(* Logix 5000 project; controller PLC_MCC1300_75F1 vendor 1 type 14 code 166 rev 32.11; software revision 32.04; part 2 of 83 *)

TYPE MAC_Popup_ZC_ALM :
STRUCT
   rgxStoppingFault : DINT[1];   // Generic stopping faults
   rgxFault : DINT[1];   // Generic faults
   rgxWarning : DINT[1];   // Generic warning
   rgxStoppingFault_M : DINT[1];   // Motor stopping faults
   rgxFault_M : DINT[1];   // Motor faults
   rgxWarning_M : DINT[1];   // Motor warning
   rgdFaultCode_M : DINT[1];   // Motor fault codes
END_STRUCT
END_TYPE

TYPE MAC_Popup_ZC_HMR :
STRUCT
   xHighPosition : BOOL;   // Popup in high position {x|x|x|x|O}
   xLowPosition : BOOL;   // Popup in low position {x|x|x|x|O}
   xPopUpCleaningEnabled : BOOL;   // Cleaning enabled on Popup
   rgdState : DINT;   // State (1=No anomaly, 3=Run, 7=Anomaly) {x|x|x|x|O}
   rgxMan : DINT;   // Manual commands {x|x|x|x|O}
END_STRUCT
END_TYPE

TYPE MAC_Popup_ZC_HMW :
STRUCT
   xLocalCleaningRequest : BOOL;   // Local cleaning popup request {x|x|x|x|O}
   xEnableDisableManualCommand : BOOL;   // Enable/disable manual command {x|x|x|x|O}
   dConvoyOffset_cmm : DINT;   // Positioning offset used for convoy positioning towards center of conveyor [mm/100] {mm/100|mm|-300|300|O}
   dSingleCapOffset_cmm : DINT;   // Positioning offset used for single cap positioning towards start of conveyor [mm/100] {mm/100|mm|-300|300|O}
   dGlassPosFromStart_cmm : DINT;   // Position of glass from start of conveyor [mm/100] {mm/100|mm|0|500|O}
   dGlassPosFromEnd_cmm : DINT;   // Position of glass from end of conveyor [mm/100] {mm/100|mm|0|500|O}
   dConvoySidePosForCenterSheet : DINT;   // Position of center sheet within 3 pieces convoy [0=left, 1=center, 2=right] {x|x|x|x|O}
   dConvoyGapForCenterSheet : DINT;   // Gap of center sheet towards selected side sheet {mm/100|mm|150|500|O}
   rgxMan : DINT;   // Manual commands {x|x|x|x|O}
   dSaturationSelection : DINT;   // Selection conveyor to start saturation {x|x|x|x|O}
END_STRUCT
END_TYPE

TYPE MAC_Popup_ZC_IN_MOTION :
STRUCT
   DR_MAJ_M : MOTION_INSTRUCTION[1];   // Drive jog
   DR_MAM_M : MOTION_INSTRUCTION[1];   // Drive positioning
   DR_MRP_M : MOTION_INSTRUCTION[1];   // Drive reset count
   DR_MAS_M : MOTION_INSTRUCTION[1];   // Drive stop
END_STRUCT
END_TYPE

TYPE MAC_Popup_ZC_OUT_MOTION :
STRUCT
   DR_MSO_M : MOTION_INSTRUCTION[1];   // Drive ON
   DR_MSF_M : MOTION_INSTRUCTION[1];   // Drive OFF
   DR_MASR_M : MOTION_INSTRUCTION[1];   // Drive reset faults
   DR_MAJ_M : MOTION_INSTRUCTION[1];   // Drive jog
   DR_MAM_M : MOTION_INSTRUCTION[1];   // Drive positioning
   DR_MRP_M : MOTION_INSTRUCTION[1];   // Drive reset count
   DR_MCD_M : MOTION_INSTRUCTION[1];   // Drive change speed
   DR_MAS_M : MOTION_INSTRUCTION[1];   // Drive stop
END_STRUCT
END_TYPE

TYPE MAC_Rotator :
STRUCT
   ST_xInitialConditionOK : BOOL;   // Initial condition OK
   ST_xCleaningConditionOK : BOOL;   // Cleaning condition OK
   ST_xCleaningAccepted : BOOL;   // Cleaning accepted
   ST_xReqCleaning : BOOL;   // Request cleaning
   ST_xPhasesInProgress : BOOL;   // Phases in progress
   ST_xStopMachineFault : BOOL;   // Stopped machine fault
   ST_xStopNextCycleFault : BOOL;   // Stopped next cycle fault
   ST_xConditionOKStopCycle : BOOL;   // Condition OK for stop cycle
   ST_xOutputEnable : BOOL;   // Output enable
   ST_xMachineAlarm : BOOL;   // Machine alarm
   ST_xFeedbackRotation : BOOL;   // Feedback rotation
   ST_xWaitMachineStop : BOOL;   // Wait machine stop
   ST_xEnableControlError : BOOL;   // Enable control error
   ST_xManualMode : BOOL;   // Manual mode enabled
   PH_x : DINT;   // Phases
   INPUT_rRotatorPosition_cdeg : REAL;   // Rotator actual angle position [°/100]
   INPUT_xBrakingResistor : BOOL;   // Braking resistor
   INPUT_xConditionToDescent : BOOL;   // Condition OK for descent
   INPUT_xDriveError : BOOL;   // Drive error
   INPUT_xDriveFeedback : BOOL;   // Drive feedback
   INPUT_xFeedbackLifting : BOOL;   // Feedback lifting
   INPUT_xHighPosition : BOOL;   // High position
   INPUT_xLowPosition : BOOL;   // Low position
   INPUT_xLocalSafetySwitchLifting : BOOL;   // Local safety switch lifting
   INPUT_xLocalSafetySwitchRotation : BOOL;   // Local safety switch rotation
   INPUT_xMotorThermalProbe : BOOL;   // Motor thermal probe
   INPUT_xProtectionMotorLifting : BOOL;   // Protection motor lifting
   INPUT_xProtectionMotorRotation : BOOL;   // Protection motor rotation
   INPUT_xDriveInhibit : BOOL;   // Drive inhibit
   INPUT_xDriveReady : BOOL;   // Drive ready
   OUTPUT_xBrakeRelease : BOOL;   // Brake release
   OUTPUT_xDescent : BOOL;   // Descent frame
   OUTPUT_xDriveEnable : BOOL;   // Drive enable
   OUTPUT_xJog : BOOL;   // Jog mode
   OUTPUT_xReverse : BOOL;   // Counterclockwise rotation
   OUTPUT_xRise : BOOL;   // Rise frame
   OUTPUT_xRun : BOOL;   // Clockwise rotation
   AUX_dDistanceCenter_cmm : DINT;   // Distance split line from center rotator frame [mm/10] (#COSTANT#)
   AUX_rTotalWeight_kg : REAL;   // Total weight [Kg]
   tmON_DelayFrameUP : TIMER;
   tmON_DelayRotatorInRun : TIMER;
   tmOF_DriveEnable : TIMER;   // Drive enable
   tmON_FeedbackTimeOutLifting : TIMER;   // Feedback time out lifting
   tmON_FeedbackTimeOutRotation : TIMER;   // Feedback time out rotation
   tmON_FramePosError : TIMER;   // Frame lifting position error
   tmON_RotatePosError : TIMER;   // Rotate positioning error
   tmON_PresetEncoder : TIMER;   // Preset ecoder
   tmON_DelayBrakeON : TIMER;   // Delay brake ON
END_STRUCT
END_TYPE

TYPE MAC_Rotator_ALM :
STRUCT
   rgxStoppingFault : DINT[1];   // Generic stopping faults
   rgxFault : DINT[1];   // Generic faults
   rgxWarning : DINT[1];   // Generic warning
   rgxStoppingFault_M : DINT[1];   // Motor stopping faults
   rgxFault_M : DINT[1];   // Motor faults
   rgxWarning_M : DINT[1];   // Motor warning
   rgdFaultCode_M : DINT[1];   // Motor fault codes
END_STRUCT
END_TYPE

TYPE MAC_Rotator_HMR :
STRUCT
   xHighPosition : BOOL;   // Rotator in high position {x|x|x|x|O}
   xLowPosition : BOOL;   // Rotator in low position {x|x|x|x|O}
   dState : DINT;   // State (1=No anomaly, 3=Run, 7=Anomaly) {x|x|x|x|O}
   dActualAngle_cdeg : DINT;   // Rotator actual angle position [°/100] {deg/100|deg|x|x|O}
   rgxMan : DINT;   // Manual commands {x|x|x|x|O}
END_STRUCT
END_TYPE

TYPE MAC_Rotator_HMW :
STRUCT
   xPresetEnc : BOOL;   // Preset encoder rotator {x|x|x|x|O}
   dLowSpeed_deg_s : DINT;   // Low speed rotator [°/s] {deg/s|deg/s|x|x|O}
   dLowRamp_deg_s2 : DINT;   // Low ramps rotator [°/s2] {deg/s2|deg/s2|x|x|O}
   dHighSpeed_deg_s : DINT;   // High speed rotator [°/s] {deg/s|deg/s|x|x|O}
   dHighRamp_deg_s2 : DINT;   // High ramps rotator [°/s2] {deg/s2|deg/s2|x|x|O}
   dJogSpeed_deg_s : DINT;   // Jog speed rotator [°/s] {deg/s|deg/s|x|x|O}
   rgxMan : DINT;   // Manual commands {x|x|x|x|O}
END_STRUCT
END_TYPE

TYPE MAC_SafetyAccess :
STRUCT
   xMxx0S_ConditionOK : BOOL;   // Mxx0S.Condition ok for request access area
   xMxx0S_SafetyOK : BOOL;   // Mxx0S.Area safety ok
   xMxx1S_ConditionOK : BOOL;   // Mxx1S.Condition ok for request access area
   xMxx1S_SafetyOK : BOOL;   // Mxx1S.Area safety ok
END_STRUCT
END_TYPE

TYPE MAC_SafetyAccess_ALM :
STRUCT
   rgxFault : DINT[2];   // Faults
END_STRUCT
END_TYPE

TYPE MAC_SafetyAccess_HMR :
STRUCT
   iMxx0S_State : DINT;   // Mxx0S.State (1=ok, 2=Access request, 4=Access done, 8=Request accepted) {x|x|x|x|O}
   iMxx1S_State : DINT;   // Mxx1S.State (1=ok, 2=Access request, 4=Access done, 8=Request accepted) {x|x|x|x|O}
END_STRUCT
END_TYPE

TYPE MAC_SpeedUp :
STRUCT
   ST_xConditionOKForSQC : BOOL;   // Condition OK for SQC plate
   ST_xConditionOKForConvoy : BOOL;   // Condition OK for convoy creation
   ST_xConditionOKChangeSpeed : BOOL;   // Condition OK for change speed
   ST_xCapDimensionOK : BOOL;   // Snapped cap dimension OK
   ST_xLastPlateInConvoy : BOOL;   // Last plate in convoy
   ST_xFirstGlassAfterClean : BOOL;   // First glass after cleaning
   ST_xReqCulletOnMissSnap : BOOL;   // Request redirect plate to cullet on missing snap (NOT USED)
   ST_xReqCulletAfterMissSnap : BOOL;   // Request redirect to cullet the plate after missing snap (NOT USED)
   ST_xChangeThicknessActive : BOOL;   // Change thickness active
   ST_xControlSnapActive : BOOL;   // Control snap active
   ST_xSpeedInc10perc : BOOL;   // Speed increase of 10% when high thickness
   ST_xAccDecLowForThicknessHigh : BOOL;   // Slowing acceleration and deceleration for high thickness
   ST_xMemoryMissingSnap : BOOL;   // Memory of missing snap
   ST_xStopMachineFault : BOOL;   // Stop for machine fault
   ST_xStopNextCycleFault : BOOL;   // Stop next cycle for fault
   ST_xWarningFault : BOOL;   // Warning fault
   ST_xPlateComing : BOOL;   // Plate coming from previous conveyor
   ST_xGapCreation : BOOL;   // Gap creation
   OSR_xNewData : BOOL;   // OSR New data
   OSR_xSnapDone : BOOL;   // OSR Snap done
   OSR_xControlSnapOK : BOOL;   // OSR Control snap OK
   OSR_xMissingSnap : BOOL;   // OSR Missing snap
   OSR_xResetDimensionZ200 : BOOL;   // OSR Reset dimension Z200
   OSR_xAccDecLowForThicknessHigh : BOOL;   // OSR Slowing acceleration and deceleration for high thickness
   OSR_xAccDecHighForThicknessLow : BOOL;   // OSR Increasing acceleration and deceleration for low thickness
   OS_xNewData : BOOL;   // OS New data
   OS_xSnapDone : BOOL;   // OS Snap done
   OS_xControlSnapOK : BOOL;   // OS Control snap OK
   OS_xMissingSnap : BOOL;   // OS Missing snap
   OS_xWrongDimension : BOOL;   // OS Wrong dimension
   OS_xLastPlateMissingSnap : BOOL;   // OS Last plate missing snap
   OS_xAccDecLowForThicknessHigh : BOOL;   // OS Slowing acceleration and deceleration for high thickness
   OS_xAccDecHighForThicknessLow : BOOL;   // OS Increasing acceleration and deceleration for low thickness
   OS_xChangeAccDec : BOOL;   // OS Change acceleration and deceleration
   INPUT_xSnapDoneHW : BOOL;   // Snap done signal on hardware
   INPUT_xControlSnap1 : BOOL;   // Control snap photocell 1
   INPUT_xControlSnap2 : BOOL;   // Control snap photocell 2
   INPUT_rRealSpeedInAcc_mm_min : REAL;   // Real speed in accelerating [mm/min]
   INPUT_dDecRamp_m_s2 : REAL;   // Deceleration ramp [m/s2]
   AUX_dMaxMissSnap : DINT;   // Maximum number of missing snap
   AUX_dMaxCapLength_cmm : DINT;   // Maximum cap length accepted [mm/100]
   AUX_dControlSnapLimit_cmm : DINT;   // Control snap photocell position [mm/100]
   AUX_dConveyorLength_cmm : DINT;   // Speed up conveyor length [mm/100]
   AUX_dLastDataReceived : DINT;   // LastDataReceived
   AUX_dDataSync : DINT;   // Data from Z200 synchronized [1=Data copy available)
   AUX_dNumCapConvoy : DINT;   // Number caps in convoy
   AUX_dDimensionCapCreation_cmm : DINT;   // Dimension cap still not snapped [mm/100]
   AUX_dDimensionCapMissSnap_cmm : DINT;   // Dimension cap on missing snap [mm/100]
   AUX_dNumMissSnap : DINT;   // Number of missing snap
   AUX_dDeltaSpeed_mm_min : DINT;   // Delta speed [mm/min]
   AUX_dDecSpace_cmm : DINT;   // Deceleration space [mm/100]
   AUX_dReqGapOnLastSnap_cmm : DINT;   // Request gap on last snap [mm/100]
   AUX_dConGapSetpoint_cmm : DINT;   // Convoy gap setpoint [mm/100]
   AUX_dSnapOffset_cmm : DINT;   // Snap offset [mm/100]
   AUX_dLastIndexTailSnap : DINT;   // Last snap index tail of convoy
   AUX_dFirstIndexHeadSnap : DINT;   // First snap index head of convoy
   AUX_dLastIndexMissingSnap : DINT;   // Last missing snap index
   AUX_dConvoyLengthComing : DINT;   // Convoy length coming [mm/100]
   AUX_dAccTimeForGap_ms : DINT;   // Accelaration time for gap [ms]
   AUX_dLastConvoyTailPos_cmm : DINT;   // Last convoy tail position after snap
   AUX_dGeneratingConvoyDestination : DINT;   // Destination of convoy in generation
   AUX_dConvoyIndexToAddGap : DINT;   // Convoy cap index where has to be added gap for asymmetric convoy
   AUX_dConvoyGapToAdd_cmm : DINT;   // Convoy gap to add in case of asymmetric convoy [mm/100]
   AUX_dConvoyGlassLength_cmm : DINT;   // Convoy length coming from Z200 (without gaps) [mm/100]
   AUX_dMaxConvoyLength_cmm : DINT;   // Convoy max length acceptable [mm/100]
   AUX_dSymmetricGap_cmm : DINT;   // Convoy symmetric Gap [mm/10]
   AUX_dConvoyLengthTarget_cmm : DINT;   // Convoy length target (with gaps) [mm/100]
   AUX_dNumCapsInConvoy : DINT;   // Number of caps in convoy
   AUX_dGapFromStartOfConvoy_cmm : DINT;   // Gap from start of convoy (lehr side manual sidelegs) [mm/100]
   AUX_dGapFromEndOfConvoy_cmm : DINT;   // Gap from end of convoy (breaker side manual sidelegs) [mm/100]
   AUX_dManualSideLegWidth_cmm : DINT;   // Manual side legs conveyors width [mm/100]
   AUX_dSumOfGapsInConvoy_cmm : DINT;   // Sum of all gap spaces in convoy [mm/100]
   AUX_dStandardGap_cmm : DINT;   // Standard gap space between caps [mm/100]
   rgxReqAcc : DINT;   // Requested accelerations
   xReqAccAll : BOOL;   // Request acceleration all
   AUX_rLehrStepInc_cmm : REAL;   // Lehr space increment on each scan [mm/100]
   tmON_TimeControlSnap : TIMER[2];   // Time out on control snap photocell
   tmON_GapCount : TIMER;   // Time for gap generation
   tmON_AllowStopCleaning : TIMER;   // Time for allow stop cleaning
   tSearchPlate : GP_TrackingSearchPlate_STC;   // Tracking search plate
END_STRUCT
END_TYPE

TYPE MAC_SpeedUp_ALM :
STRUCT
   rgxStoppingFault : DINT;   // Generic stopping faults
   rgxFault : DINT;   // Generic faults
   rgxWarning : DINT;   // Generic warning
END_STRUCT
END_TYPE

TYPE MAC_SpeedUp_HMR :
STRUCT
   xControlSnap1 : BOOL;   // Control snap photocell 1 {x|x|x|x|O}
   xControlSnap2 : BOOL;   // Control snap photocell 2 {x|x|x|x|O}
   dControlSnapEnabled : BOOL;   // Control snap enabled {x|x|x|x|O}
   rgdStateSensor : DINT[2];   // Control snap photocell state {x|x|x|x|O}
END_STRUCT
END_TYPE

TYPE MAC_SpeedUp_HMW :
STRUCT
   xEnableControlSnap : BOOL;   // Enable control snap {x|x|x|x|O}
   xDisableControlSnap : BOOL;   // Disable control snap {x|x|x|x|O}
END_STRUCT
END_TYPE

TYPE MAC_TrimmingDeck :
STRUCT
   CONF_dTolerance_cmm : DINT;   // Tolerance position trimming deck [mm/100]
   CONF_dStopCam_cmm : DINT;   // Stop cam position trimming deck [mm/100]
   CONF_dSlowDown_cmm : DINT;   // Slow down position trimming deck [mm/100]
   CONF_dStartPositionFrame : DINT;   // Distance from the beggining (From origin to split line) [mm/100]
   CONF_dConveyorLength_cmm : DINT;   // Conveyor length [mm/100]
   CONF_dStopPositionFrame_cmm : DINT;   // Distance of end machine from the beggining (From origin to split line) [mm/100]
   CONF_dMaxTimeToReachPosition_ms : DINT;   // Maximum time to end positioning [ms]
   CONF_dTrimDeckPreset : DINT[2];   // Trimming deck preset encoder [pulse]
   CONF_rTrimDeckPresetScaling : REAL[2];   // Trimming deck preset scaling [(mm/100) / pulse]
   CONF_dTrimDeckPresetZero_cmm : DINT[2];   // Trimming deck encoder value in zero position [mm/100]
   CONF_dTrimDeckTargetWindow_cmm : DINT[2];   // Trimming deck tollerance window on request position [mm/100]
   CONF_dTrimDeckDecWindow_cmm : DINT[2];   // Trimming deck tollerance window on deceleration position [mm/100]
   CONF_dTrimDeckCleanPos_cmm : DINT[2];   // Trimming deck cleaning position [mm/100]
   CONF_dTrimDeckMinPos_cmm : DINT[2];   // Trimming deck minimum position [mm/100]
   CONF_dTrimDeckMaxPos_cmm : DINT[2];   // Trimming deck maximum position [mm/100]
   CONF_dTrimDeckWheelsDist_cmm : DINT[2];   // Trimming deck distance from wheels support beam [mm/100]
   CONF_dTrimDeckMinRange_cmm : DINT;   // Trimming deck minimum work range [mm/100]
   CONF_dTrimDeckMaxRange_cmm : DINT;   // Trimming deck maximum work range [mm/100]
   CONF_dTrimDeckMovePos_cmm : DINT;   // Trimming deck position to start moving [mm/100]
   CONF_dTrimDeckEndArmPos_cmm : DINT;   // Trimming deck position for arming end [mm/100]
   CONF_dAutoSpeed_mm_min : DINT;   // Nominal speed in automatic mode [mm/min]
   CONF_dSlowDownSpeed_mm_min : DINT;   // Fine speed to end positioning [mm/min]
   CONF_dManualSpeed_mm_min : DINT;   // Manual speed [mm/min]
   CONF_rAcceleration_m_s2 : REAL[2];   // Trimming deck acceleration ramp [m/s2]
   CONF_rDeceleration_m_s2 : REAL[2];   // Trimming deck deceleration ramp [m/s2]
   ST_xInitialConditionOK : BOOL;   // Initial condition OK
   ST_xPhasesInProgressOpSide : BOOL;   // Phases in progress operator side
   ST_xPhasesInProgressOppOpSide : BOOL;   // Phases in progress opposite operator side
   ST_xCleaningConditionOK : BOOL;   // Cleaning condition OK
   ST_xStopMachineFault : BOOL;   // Stopped machine faults
   ST_xStopNextCycleFault : BOOL;   // Stopped next cycle faults
   ST_xConditionOKStopCycle : BOOL;   // Condition OK for stop cycle
   ST_xOutputEnable : BOOL;   // Output enable
   ST_xMachineFault : BOOL;   // Machine with faults
   ST_xWarningFault : BOOL;   // Machine with warnings
   ST_xSafetyMovement : BOOL;   // Safety movement
   ST_xHeadPresence : BOOL;   // Head presence on conveyor
   ST_xTailPresence : BOOL;   // Tail presence on conveyor
   ST_xEnableControlError : BOOL;   // Enable control error
   ST_xDoubleSizeProduction : BOOL;   // Different production size in progress
   ST_xJumboInProgress : BOOL;   // Jumbo plate in progress
   ST_xConvoyInProgress : BOOL;   // Convoy in progress
   ST_xFirstCapInConv : BOOL;   // First plate in convoy
   ST_xQualityInProgress : BOOL;   // Quality plate in progress
   ST_xCulletInProgress : BOOL;   // Cullet plate in progress
   ST_xShortestInProgress : BOOL;   // Shortest size in progress
   ST_xBiggestInProgress : BOOL;   // Biggest size in progress
   ST_xTrimDeckInWorkOpSide : BOOL;   // Trimming deck in work operator side
   ST_xTrimDeckInWorkOppOpSide : BOOL;   // Trimming deck in work opposite operator side
   ST_xCulletEdgeEnabled : BOOL;   // Trimming deck enabled for cullet edges
   ST_xInPositionOpSide : BOOL;   // Operator side frame in position
   ST_xInPositionOppOpSide : BOOL;   // Opposite operator side frame in position
   ST_xInSlowDownOpSide : BOOL;   // Operator side frame in slow down
   ST_xInSlowDownOppOpSide : BOOL;   // Opposite operator side frame in slow down
   ST_xStopCamPositionOpSide : BOOL;   // Operator side frame in stop cam position
   ST_xStopCamPositionOppOpSide : BOOL;   // Opposite operator side frame in stop cam position
   ST_xInSlowDownManualOpSide : BOOL;   // Operator side frame in manual slow down
   ST_xInSlowDownManualOppOpSide : BOOL;   // Opposite operator side frame in manual slow down
   ST_xInSlowDownManualPosOpSide : BOOL;   // Operator side frame in manual positioning slow down
   ST_xInSlowDownManualPosOppOpSide : BOOL;   // Opposite operator side frame in manual positioning slow down
   ST_xStopCamManualOpSide : BOOL;   // Operator side frame in manual stop cam
   ST_xStopCamManualOppOpSide : BOOL;   // Opposite operator side frame in manual stop cam
   ST_xStopCamManualPositionOpSide : BOOL;   // Operator side frame in manual stop cam positioning
   ST_xStopCamManualPositionOppOpSide : BOOL;   // Opposite operator side frame in manual stop cam positioning
   ST_xPositionReachedOpSide : BOOL;   // Operator side frame position reached
   ST_xPositionReachedOppOpSide : BOOL;   // Opposite operator side frame position reached
   ST_xInitialConditionHomeOpSide : BOOL;   // Initial condition for home cycle operator side
   ST_xInitialConditionHomeOppOpSide : BOOL;   // Initial condition for home cycle opposite operator side
   ST_xAxleHomedOpSide : BOOL;   // Axle homed operator side
   ST_xAxleHomedOppOpSide : BOOL;   // Axle homed opposite operator side
   ST_xReqStartMovement : BOOL;   // Request start movement
   ST_xReqAbortMovement : BOOL;   // Request abort movement
   ST_xReqResetOffset : BOOL;   // Request reset offset
   ST_xReqUpdateTarget : BOOL;   // Request update target
   OSR_xPresetEncoderOpSide : BOOL;   // OSR Preset encoder operator side
   OSR_xPresetEncoderOppOpSide : BOOL;   // OSR Preset encoder opposite operator side
   OSR_xControlWidthAuto : BOOL;   // OSR Control cap width in automatic
   OSR_xOpSideToExternal : BOOL;   // OSR Operator side to external
   OSR_xOpSideToInternal : BOOL;   // OSR Operator side to internal
   OSR_xOppOpSideToExternal : BOOL;   // OSR Opposite operator side to external
   OSR_xOppOpSideToInternal : BOOL;   // OSR Opposite operator side to internall
   OSR_xBothSideToOpSide : BOOL;   // OSR Both sides to operator side
   OSR_xBothSideToOppOpSide : BOOL;   // OSR Both sides to opposite operator side
   OSR_xStartMoveFromEth1 : BOOL;   // OSR Start moving trimming deck
   OSR_xStartMoveFromTracking : BOOL;   // OSR Start moving trimming deck
   OSR_xStartPositioning : BOOL;   // OSR Start positioning
   OSR_xUpdateTarget : BOOL;   // OSR Update target
   OSR_xReqHomeCycleOpSide : BOOL;   // OSR Request home cycle operator side
   OSR_xReqHomeCycleOppOpSide : BOOL;   // OSR Request home cycle opposite operator side
   OS_xPresetEncoderOpSide : BOOL;   // OS Preset encoder operator side
   OS_xPresetEncoderOppOpSide : BOOL;   // OS Preset encoder opposite operator side
   OS_xControlWidthAuto : BOOL;   // OS Control cap width in automatic
   OS_xStartMoveFromEth1 : BOOL;   // OS Start moving trimming deck
   OS_xStartMoveFromTracking : BOOL;   // OS Start moving trimming deck
   OS_xStartPositioning : BOOL;   // OS Start positioning
   OS_xUpdateTarget : BOOL;   // OS Update target
   OS_xReqHomeCycleOpSide : BOOL;   // OS Request home cycle operator side
   OS_xReqHomeCycleOppOpSide : BOOL;   // OS Request home cycle opposite operator side
   PH_xRequestPositionOpSide : BOOL;   // PH Request position operator side
   PH_xEndPositionOpSide : BOOL;   // PH End position operator side
   PH_xReleaseSensorHomeOpSide : BOOL;   // PH Release sensor home operaor side
   PH_xHomeCycleOpSide : BOOL;   // PH Home cycle operator side
   PH_xEndHomeCycleOpSide : BOOL;   // PH End Home cycle operator side
   PH_xRequestPositionOppOpSide : BOOL;   // PH Request position opposite operator side
   PH_xEndPositionOppOpSide : BOOL;   // PH End position opposite operator side
   PH_xReleaseSensorHomeOppOpSide : BOOL;   // PH Release sensor home opposite operaor side
   PH_xHomeCycleOppOpSide : BOOL;   // PH Home cycle opposite operator side
   PH_xEndHomeCycleOppOpSide : BOOL;   // PH End Home cycle opposite operator side
   INPUT_xSBControlWidthAuto : BOOL;   // Control cap width in automatic
   INPUT_xSQAntiCollision : BOOL;   // Anti collision sensor
   INPUT_xFrameInOpSidePosition : DINT;   // Frame in operator side position
   INPUT_xFrameInOppOpSidePosition : DINT;   // Frame in opposite operator side position
   INPUT_xBrakingResistor : DINT;   // Braking Resistor
   INPUT_xDriveInhibit : DINT;   // Drive inhibit
   INPUT_xDriveReady : DINT;   // Drive ready
   INPUT_xDriveError : DINT;   // Drive Error
   INPUT_xDriveFeedback : DINT;   // Drive Feedback
   INPUT_xDriveDeceleration : DINT;   // Drive deceleration
   INPUT_xLocalSafetySwitch : DINT;   // Local Safety Switch
   INPUT_xMotorThermalProbe : DINT;   // Motor Thermal Probe
   INPUT_xProtectionMotor : DINT;   // Protection Motor
   INPUT_xOverstrokeExternal : DINT;   // External overstroke
   INPUT_xDriveHomedStatus : DINT;   // Drive homed status
   INPUT_xSQTrimDeckExternalStop : DINT;   // Trimming deck to stop external position
   INPUT_xSQTrimDeckInternalStop : DINT;   // Trimming deck to stop internal position
   INPUT_xSATrimDeckToExternal : DINT;   // Trimming deck selector to external side
   INPUT_xSATrimDeckToInternal : DINT;   // Trimming deck selector to internal side
   INPUT_xSATrimDeckToOpSide : DINT;   // Trimming deck selector to operator side
   INPUT_xSATrimDeckToOppOpSide : DINT;   // Trimming deck selector to opposite operator side
   INPUT_dEncoderPulse : DINT[2];   // Trimming deck encoder [pulse]
   OUTPUT_xSBControlWidthAuto : BOOL;   // Control cap width in automatic
   OUTPUT_xDriveReset : DINT;   // Drive reset faults
   OUTPUT_xDriveEnable : DINT;   // Output
   OUTPUT_xRun : DINT;   // Run
   OUTPUT_xReverse : DINT;   // Reverse
   OUTPUT_xPositioning : DINT;   // Positioning
   OUTPUT_xHoming : DINT;   // Homing
   OUTPUT_xChangeSpeed : DINT;   // Change speed
   OUTPUT_dEncoder : DINT;   // Encoder
   OUTPUT_xSATrimDeckToExternal : DINT;   // Trimming deck selector to external side
   OUTPUT_xSATrimDeckToInternal : DINT;   // Trimming deck selector to internal side
   OUTPUT_xSATrimDeckToOpSide : DINT;   // Trimming deck selector to operator side
   OUTPUT_xSATrimDeckToOppOpSide : DINT;   // Trimming deck selector to opposite operator side
   AUX_dHeadPosition_cmm : DINT;   // Plate head position [mm/100]
   AUX_dTailPosition_cmm : DINT;   // Plate tail position [mm/100]
   AUX_dReqTargetPos_cmm : DINT[2];   // Request target position [mm/100]
   AUX_dOffset_cmm : DINT[2];   // Offset position [mm/100]
   AUX_dTarget_cmm : DINT[2];   // Trimming deck target position without offset [mm/100]
   AUX_dFinalTarget_cmm : DINT[2];   // Trimming deck final target position [mm/100]
   AUX_dActTransPosition_cmm : DINT[2];   // Actual translation position [mm/100]
   AUX_dCopyEncoderValue_cmm : DINT[2];   // Copy encoder value [mm/100]
   AUX_dCounterForAlarmEnc_cmm : DINT[2];   // Counter for encoder alarm [mm/100]
   AUX_dReqSpeed_mm_min : DINT[2];   // Trimming deck requested speed [mm/min]
   AUX_dRealSpeed_mm_min : DINT[2];   // Trimming deck real speed [mm/min]
   AUX_dPositionStartAnyway_cmm : DINT;   // Start anyway position [mm/100]
   AUX_tSearchPlateData : UDT_SearchPlateAuxData;   // Auxiliary data for searching plate
   tmON_RequestHomeCycle : TIMER[2];   // Request home cycle
   tmON_EncPreset : TIMER[2];   // Encoder preset
   tmON_CheckEncoderTimeOut : TIMER[2];   // Check encoder time out
   tmON_FeedbackTimeOut : TIMER[2];   // Feedback time out
   tmOF_DriveEnable : TIMER[2];   // Drive enable timer
   tmOF_DelayOnChangeDirection : TIMER[4];   // Delay on change direction
   tmON_FeedbackDriveReady : TIMER[2];   // Drive ready feedback timer
   tmON_ReadyToMoveDelay : TIMER[2];   // Drive ready to move timer
   tmON_Wait : TIMER;   // Wait for glass process
END_STRUCT
END_TYPE

TYPE MAC_TrimmingDeck_ALM :
STRUCT
   rgxStoppingFault : MAC_TrimmingDeck_ALM_SF[1];   // Generic stopping faults
   rgxFault : MAC_TrimmingDeck_ALM_F[1];   // Generic faults
   rgxWarning : MAC_TrimmingDeck_ALM_W[1];   // Generic warning
   rgxStoppingFault_M : MAC_TrimmingDeck_ALM_SFM[2];   // Motor stopping faults
   rgxFault_M : MAC_TrimmingDeck_ALM_FM[2];   // Motor faults
   rgxWarning_M : MAC_TrimmingDeck_ALM_WM[2];   // Motor warning
   rgdFaultCode_M : DINT[2];   // Motor fault codes
END_STRUCT
END_TYPE

TYPE MAC_TrimmingDeck_ALM_F :
STRUCT
   x0 : BOOL;   // Anticollision frame sensor
   x1 : BOOL;
   x2 : BOOL;
   x3 : BOOL;
   x4 : BOOL;
   x5 : BOOL;
   x6 : BOOL;
   x7 : BOOL;
   x8 : BOOL;
   x9 : BOOL;
   x10 : BOOL;
   x11 : BOOL;
   x12 : BOOL;
   x13 : BOOL;
   x14 : BOOL;
   x15 : BOOL;
   x16 : BOOL;
   x17 : BOOL;
   x18 : BOOL;
   x19 : BOOL;
   x20 : BOOL;
   x21 : BOOL;
   x22 : BOOL;
   x23 : BOOL;
   x24 : BOOL;
   x25 : BOOL;
   x26 : BOOL;
   x27 : BOOL;
   x28 : BOOL;
   x29 : BOOL;
   x30 : BOOL;
   x31 : BOOL;
END_STRUCT
END_TYPE

TYPE MAC_TrimmingDeck_ALM_FM :
STRUCT
   x0 : BOOL;
   x1 : BOOL;
   x2 : BOOL;
   x3 : BOOL;
   x4 : BOOL;
   x5 : BOOL;
   x6 : BOOL;
   x7 : BOOL;
   x8 : BOOL;
   x9 : BOOL;
   x10 : BOOL;
   x11 : BOOL;
   x12 : BOOL;
   x13 : BOOL;
   x14 : BOOL;
   x15 : BOOL;
   x16 : BOOL;
   x17 : BOOL;
   x18 : BOOL;
   x19 : BOOL;
   x20 : BOOL;
   x21 : BOOL;
   x22 : BOOL;
   x23 : BOOL;
   x24 : BOOL;
   x25 : BOOL;
   x26 : BOOL;
   x27 : BOOL;
   x28 : BOOL;
   x29 : BOOL;
   x30 : BOOL;
   x31 : BOOL;
END_STRUCT
END_TYPE

TYPE MAC_TrimmingDeck_ALM_SF :
STRUCT
   x0 : BOOL;
   x1 : BOOL;
   x2 : BOOL;
   x3 : BOOL;
   x4 : BOOL;
   x5 : BOOL;
   x6 : BOOL;
   x7 : BOOL;
   x8 : BOOL;
   x9 : BOOL;
   x10 : BOOL;
   x11 : BOOL;
   x12 : BOOL;
   x13 : BOOL;
   x14 : BOOL;
   x15 : BOOL;
   x16 : BOOL;
   x17 : BOOL;
   x18 : BOOL;
   x19 : BOOL;
   x20 : BOOL;
   x21 : BOOL;
   x22 : BOOL;
   x23 : BOOL;
   x24 : BOOL;
   x25 : BOOL;
   x26 : BOOL;
   x27 : BOOL;
   x28 : BOOL;
   x29 : BOOL;
   x30 : BOOL;
   x31 : BOOL;
END_STRUCT
END_TYPE

TYPE MAC_TrimmingDeck_ALM_SFM :
STRUCT
   x0 : BOOL;   // Protection motor
   x1 : BOOL;   // Drive error
   x2 : BOOL;   // Drive feedback error
   x3 : BOOL;   // Local safety switch
   x4 : BOOL;   // Motor thermal probe
   x5 : BOOL;   // Braking resistor fault
   x6 : BOOL;   // Encoder error
   x7 : BOOL;
   x8 : BOOL;
   x9 : BOOL;
   x10 : BOOL;
   x11 : BOOL;
   x12 : BOOL;
   x13 : BOOL;
   x14 : BOOL;
   x15 : BOOL;
   x16 : BOOL;
   x17 : BOOL;
   x18 : BOOL;
   x19 : BOOL;
   x20 : BOOL;
   x21 : BOOL;
   x22 : BOOL;
   x23 : BOOL;
   x24 : BOOL;
   x25 : BOOL;
   x26 : BOOL;
   x27 : BOOL;
   x28 : BOOL;
   x29 : BOOL;
   x30 : BOOL;
   x31 : BOOL;
END_STRUCT
END_TYPE

TYPE MAC_TrimmingDeck_ALM_W :
STRUCT
   x0 : BOOL;
   x1 : BOOL;
   x2 : BOOL;
   x3 : BOOL;
   x4 : BOOL;
   x5 : BOOL;
   x6 : BOOL;
   x7 : BOOL;
   x8 : BOOL;
   x9 : BOOL;
   x10 : BOOL;
   x11 : BOOL;
   x12 : BOOL;
   x13 : BOOL;
   x14 : BOOL;
   x15 : BOOL;
   x16 : BOOL;
   x17 : BOOL;
   x18 : BOOL;
   x19 : BOOL;
   x20 : BOOL;
   x21 : BOOL;
   x22 : BOOL;
   x23 : BOOL;
   x24 : BOOL;
   x25 : BOOL;
   x26 : BOOL;
   x27 : BOOL;
   x28 : BOOL;
   x29 : BOOL;
   x30 : BOOL;
   x31 : BOOL;
END_STRUCT
END_TYPE

TYPE MAC_TrimmingDeck_ALM_WM :
STRUCT
   x0 : BOOL;
   x1 : BOOL;
   x2 : BOOL;
   x3 : BOOL;
   x4 : BOOL;
   x5 : BOOL;
   x6 : BOOL;
   x7 : BOOL;
   x8 : BOOL;
   x9 : BOOL;
   x10 : BOOL;
   x11 : BOOL;
   x12 : BOOL;
   x13 : BOOL;
   x14 : BOOL;
   x15 : BOOL;
   x16 : BOOL;
   x17 : BOOL;
   x18 : BOOL;
   x19 : BOOL;
   x20 : BOOL;
   x21 : BOOL;
   x22 : BOOL;
   x23 : BOOL;
   x24 : BOOL;
   x25 : BOOL;
   x26 : BOOL;
   x27 : BOOL;
   x28 : BOOL;
   x29 : BOOL;
   x30 : BOOL;
   x31 : BOOL;
END_STRUCT
END_TYPE

TYPE MAC_TrimmingDeck_HMR :
STRUCT
   xControlWidthEnabled : BOOL;   // Control cap width in automatic enabled {x|x|x|x|O}
   xControlWanderEnabled : BOOL;   // Control cap wander in automatic enabled {x|x|x|x|O}
   xCulletEdgeEnabled : BOOL;   // Enable/Disable cullet edges trimming {x|x|x|x|O}
   xOpeningOnCleaningEnabled : BOOL;   // Opening trimming deck on cleaning mode enabled {x|x|x|x|O}
   xHooked : BOOL;   // Plate hooked {x|x|x|x|O}
   rgdState : DINT[2];   // State (1=No alarm, 3=Run, 7=Alarm) {x|x|x|x|O}
   dGrossWidthInProgress_cmm : DINT;   // Gross width in progress [mm/100] {mm/100|mm|x|x|O}
   dNetWidthInProgress_cmm : DINT;   // Net width in progress [mm/100] {mm/100|mm|x|x|O}
   dCutWanderInProgress_cmm : DINT;   // Cut wander in progress [mm/100] {mm/100|mm|x|x|O}
   rgdDEdgeWidth_cmm : DINT[2];   // Double edge width [mm/100] {mm/100|mm|x|x|O}
   rgdTarget_cmm : DINT[2];   // Trimming deck request position [mm/100] {mm/100|mm|x|x|O}
   rgdPosition_cmm : DINT[2];   // Trimming deck actual position [mm/100] {mm/100|mm|x|x|O}
   rgdOffsetEachSide_cmm : DINT[2];   // Trimming deck offset on each side [mm/100] {mm/100|mm|x|x|O}
   dOffsetBothSide_cmm : DINT;   // Trimming deck offset on both sides [mm/100] {mm/100|mm|x|x|O}
   dDistBetweenSides_cmm : DINT;   // Trimming deck distance between external conveyor wheels [mm/100] {mm/100|mm|x|x|O}
   dHead_cmm : DINT;   // Head plate position [mm/100] {mm/100|mm|x|x|O}
   dTail_cmm : DINT;   // Tail plate position [mm/100] {mm/100|mm|x|x|O}
   dWander_cmm : DINT;   // Wander plate [mm/100] {mm/100|mm|x|x|O}
   rgxMan : MAC_TrimmingDeck_HMWR_Man;   // Manual commands {x|x|x|x|O}
END_STRUCT
END_TYPE
